REGION Network 2
   "TimeServerCom"(BatchEndTime := "OPC".CON_Material.NewBatchEndTime,
                   "Date" => "PrinterData".CON.PrinterBagData."Date",
                   "Time" => "PrinterData".CON.PrinterBagData."Time",
                   BatchStatus => "OPC".CON_Material.BatchStatus);
END_REGION

REGION Network 3
   IF NOT "PrinterData".CON.PrinterSelection THEN
       #Domino(RemoteAddress := "PrinterData".CON.PrinterBagData.RemoteAddress,   // "Domino_AX"
               ConnectionStatus := #ComandsSending_Domino.connected AND #BatchSending_Domino.connected,
               ID := 2,
               ConType := True,
               ArtFlag := #HandleComBag.ActualArtFlag,
               MDR_Flag := #HandleComBag.ActualMDR_Flag,
               BatchStatus := "OPC".CON_Material.BatchStatus,
               BatchNumber := "OPC".CON_Material.ActualBatchNumber,
               ArtBaseNumber := "OPC".CON_Material.ActualArtBaseNumber,
               MarketRegCode := "OPC".CON_Material.ActualMarketRegCode,
               ExtDate := "OPC".CON_Material.ActualBBD,
               "Date" := "PrinterData".CON.PrinterBagData."Date",
               "Time" := "PrinterData".CON.PrinterBagData."Time",
               PlainDataChanged := #HandleComBag.NewDataPlain,
               DataReceived := #ComandsSending_Domino.dataReceived,
               DataReceivedBatch := #BatchSending_Domino.dataReceived,
               DataSent := #ComandsSending_Domino.sending,
               DataSentBatch := #BatchSending_Domino.sending,
               TimeSynchPeriod := "TimeSynchPeriod",
               AlarmCheckPeriod := "AlarmCheckPeriod",
               RDataBatch := "PrinterData".CON.PrinterBagData.RdataBatch,
               RData := "PrinterData".CON.PrinterBagData.RData,
               NMDR_LabelName := "PrinterData".CON.PrinterBagData.NonMDR_LabelName,
               LabelSelecting := "PrinterData".CON.PrinterBagData.Initialization,
               ErrorIP => "CON_ErrorIP",
               BatchOK => "PrinterData".CON.PrinterBagData.BatchOK,
               TimeOK => "PrinterData".CON.PrinterBagData.TimeOK);
   END_IF;
END_REGION

REGION Network 4
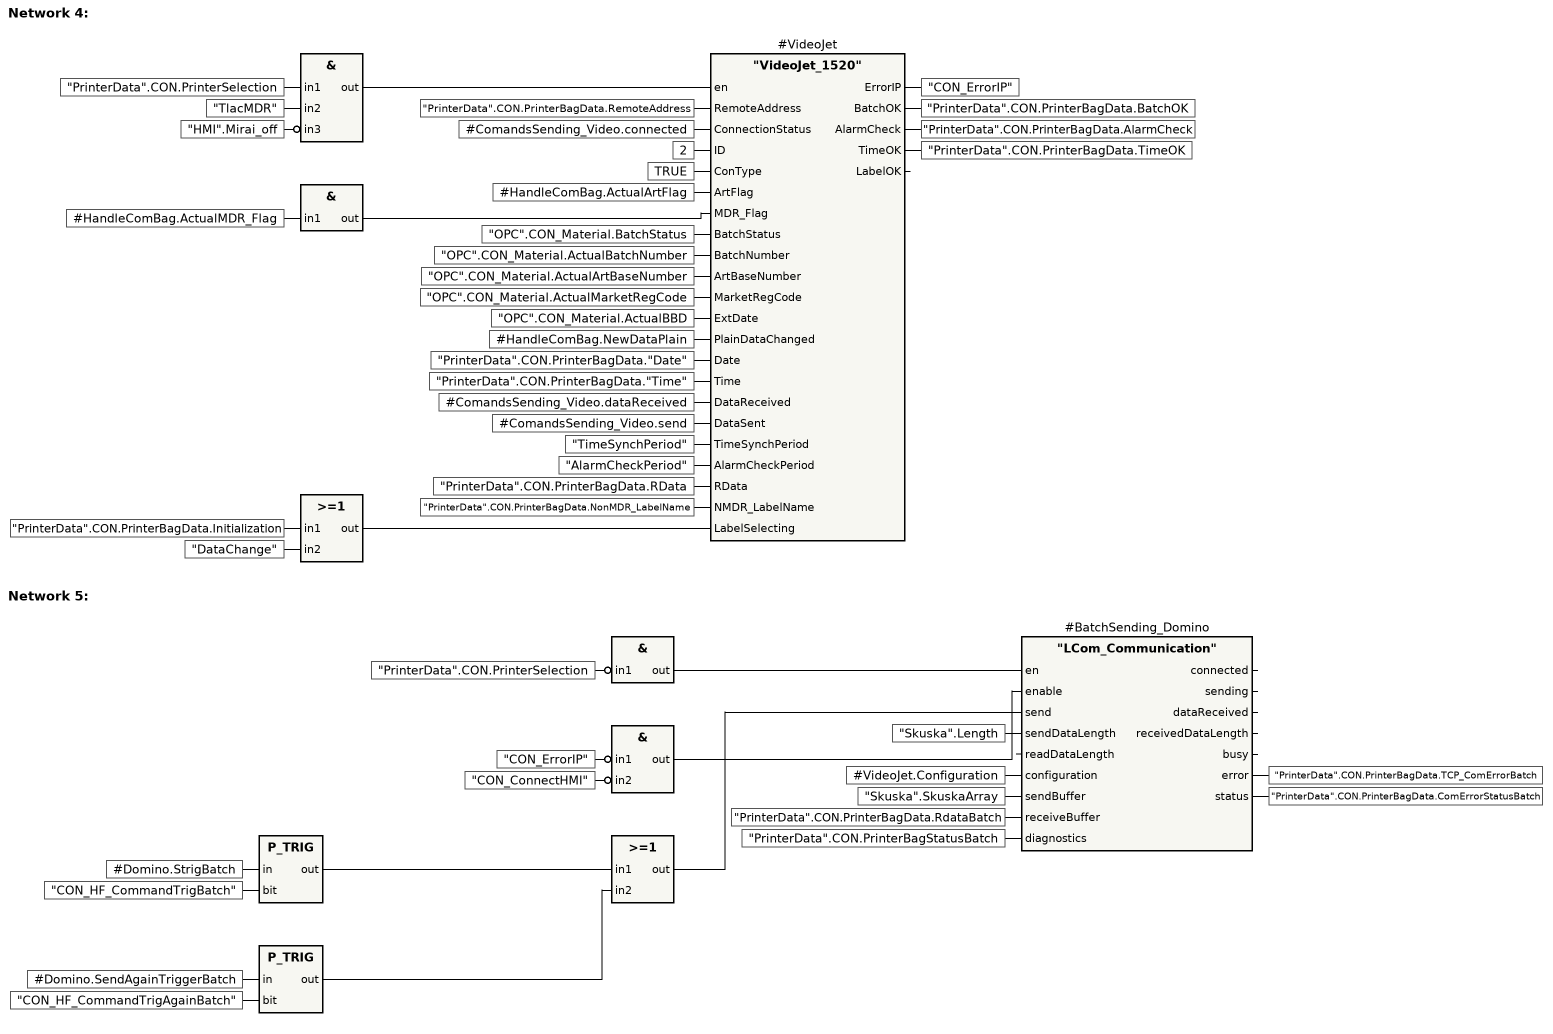
   IF "PrinterData".CON.PrinterSelection AND "TlacMDR" AND NOT "HMI".Mirai_off THEN
       #VideoJet(RemoteAddress := "PrinterData".CON.PrinterBagData.RemoteAddress,   // "VideoJet_1520"
                 ConnectionStatus := #ComandsSending_Video.connected,
                 ID := 2,
                 ConType := TRUE,
                 ArtFlag := #HandleComBag.ActualArtFlag,
                 MDR_Flag := #HandleComBag.ActualMDR_Flag,
                 BatchStatus := "OPC".CON_Material.BatchStatus,
                 BatchNumber := "OPC".CON_Material.ActualBatchNumber,
                 ArtBaseNumber := "OPC".CON_Material.ActualArtBaseNumber,
                 MarketRegCode := "OPC".CON_Material.ActualMarketRegCode,
                 ExtDate := "OPC".CON_Material.ActualBBD,
                 PlainDataChanged := #HandleComBag.NewDataPlain,
                 "Date" := "PrinterData".CON.PrinterBagData."Date",
                 "Time" := "PrinterData".CON.PrinterBagData."Time",
                 DataReceived := #ComandsSending_Video.dataReceived,
                 DataSent := #ComandsSending_Video.send,
                 TimeSynchPeriod := "TimeSynchPeriod",
                 AlarmCheckPeriod := "AlarmCheckPeriod",
                 RData := "PrinterData".CON.PrinterBagData.RData,
                 NMDR_LabelName := "PrinterData".CON.PrinterBagData.NonMDR_LabelName,
                 LabelSelecting := "PrinterData".CON.PrinterBagData.Initialization OR "DataChange",
                 ErrorIP => "CON_ErrorIP",
                 BatchOK => "PrinterData".CON.PrinterBagData.BatchOK,
                 AlarmCheck => "PrinterData".CON.PrinterBagData.AlarmCheck,
                 TimeOK => "PrinterData".CON.PrinterBagData.TimeOK);
   END_IF;
END_REGION

REGION Network 5
   #_w1 := #Domino.StrigBatch AND NOT "CON_HF_CommandTrigBatch";   // rising edge
   "CON_HF_CommandTrigBatch" := #Domino.StrigBatch;
   #_w2 := #Domino.SendAgainTriggerBatch AND NOT "CON_HF_CommandTrigAgainBatch";   // rising edge
   "CON_HF_CommandTrigAgainBatch" := #Domino.SendAgainTriggerBatch;
   IF NOT "PrinterData".CON.PrinterSelection THEN
       #BatchSending_Domino(enable := NOT "CON_ErrorIP" AND NOT "CON_ConnectHMI",   // "LCom_Communication"
                            send := #_w1 OR #_w2,
                            sendDataLength := "Skuska".Length,
                            configuration := #VideoJet.Configuration,
                            sendBuffer := "Skuska".SkuskaArray,
                            receiveBuffer := "PrinterData".CON.PrinterBagData.RdataBatch,
                            diagnostics := "PrinterData".CON.PrinterBagStatusBatch,
                            error => "PrinterData".CON.PrinterBagData.TCP_ComErrorBatch,
                            status => "PrinterData".CON.PrinterBagData.ComErrorStatusBatch);
   END_IF;
END_REGION

REGION Network 6
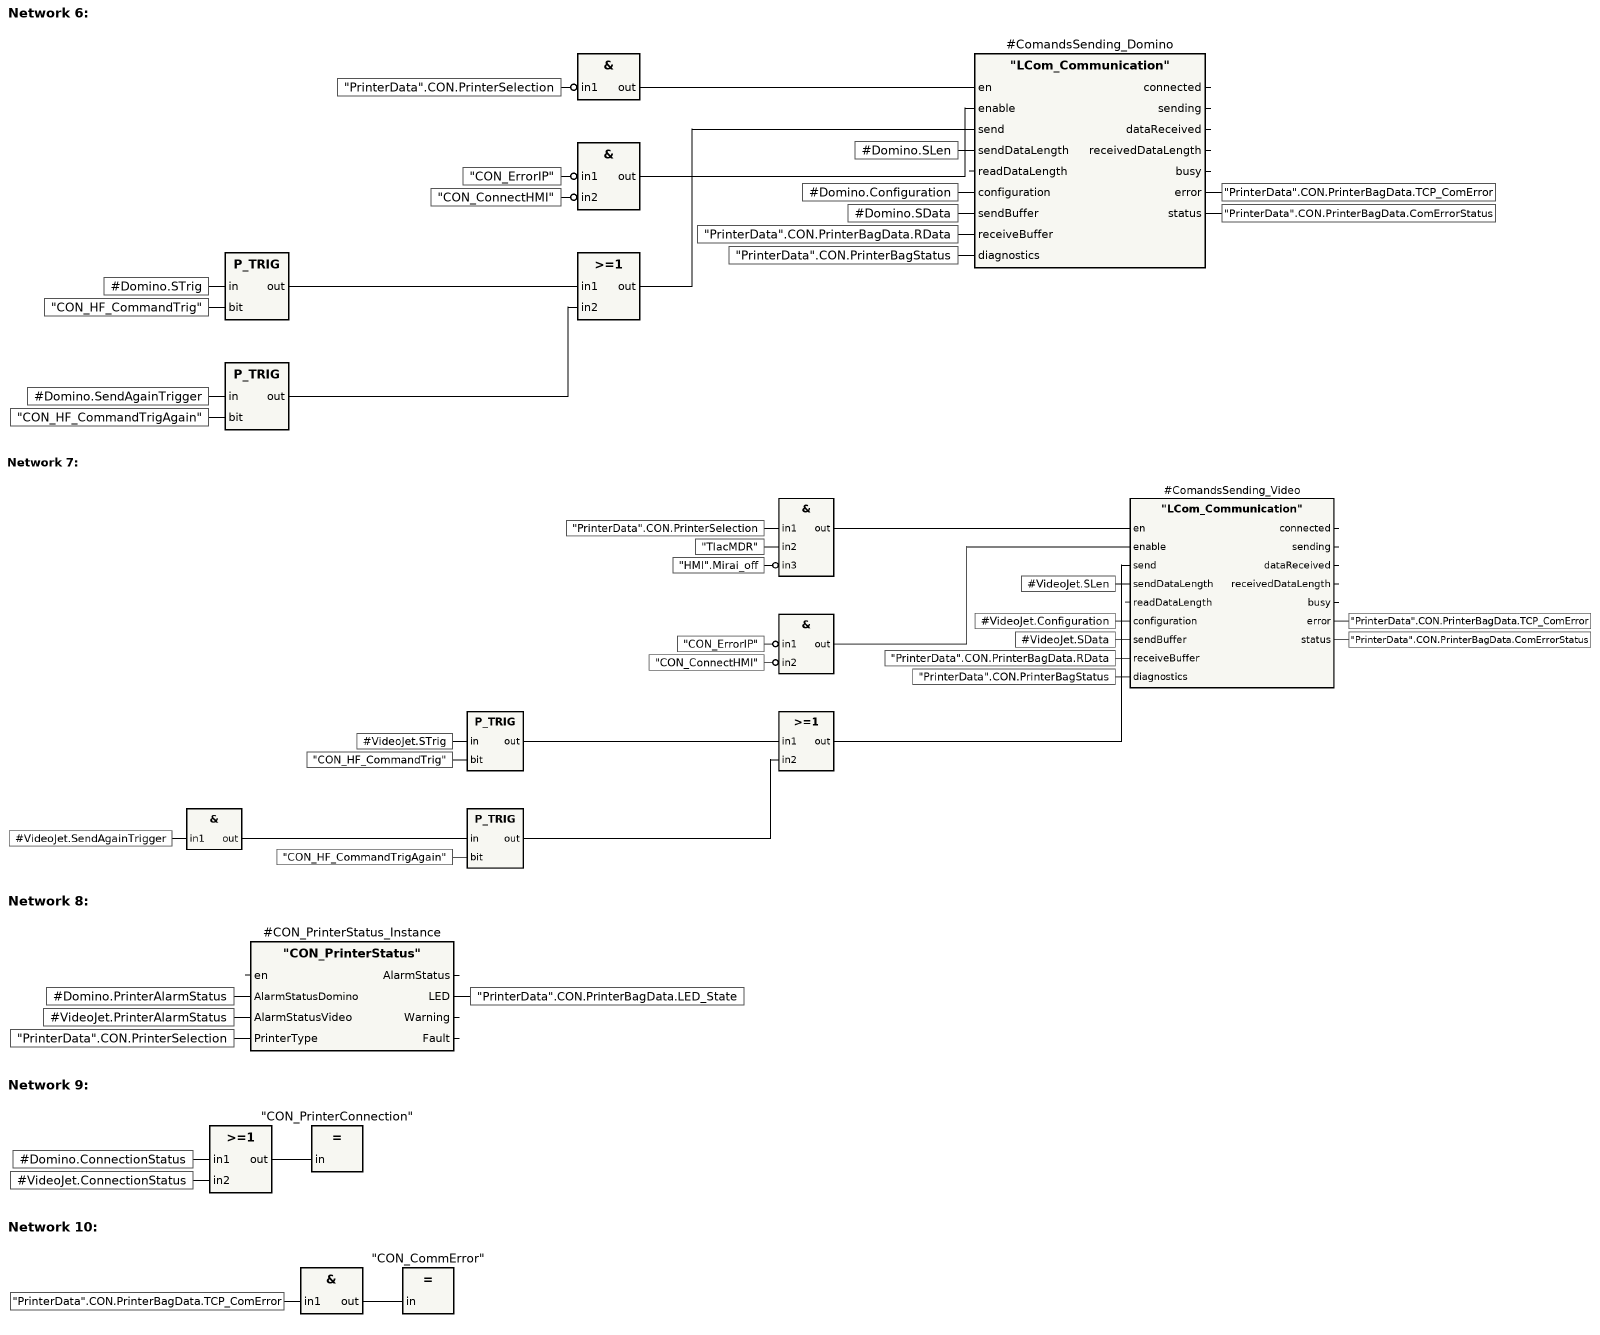
   #_w1 := #Domino.STrig AND NOT "CON_HF_CommandTrig";   // rising edge
   "CON_HF_CommandTrig" := #Domino.STrig;
   #_w2 := #Domino.SendAgainTrigger AND NOT "CON_HF_CommandTrigAgain";   // rising edge
   "CON_HF_CommandTrigAgain" := #Domino.SendAgainTrigger;
   IF NOT "PrinterData".CON.PrinterSelection THEN
       #ComandsSending_Domino(enable := NOT "CON_ErrorIP" AND NOT "CON_ConnectHMI",   // "LCom_Communication"
                              send := #_w1 OR #_w2,
                              sendDataLength := #Domino.SLen,
                              configuration := #Domino.Configuration,
                              sendBuffer := #Domino.SData,
                              receiveBuffer := "PrinterData".CON.PrinterBagData.RData,
                              diagnostics := "PrinterData".CON.PrinterBagStatus,
                              error => "PrinterData".CON.PrinterBagData.TCP_ComError,
                              status => "PrinterData".CON.PrinterBagData.ComErrorStatus);
   END_IF;
END_REGION

REGION Network 7
   #_w1 := #VideoJet.STrig AND NOT "CON_HF_CommandTrig";   // rising edge
   "CON_HF_CommandTrig" := #VideoJet.STrig;
   #_w2 := #VideoJet.SendAgainTrigger AND NOT "CON_HF_CommandTrigAgain";   // rising edge
   "CON_HF_CommandTrigAgain" := #VideoJet.SendAgainTrigger;
   IF "PrinterData".CON.PrinterSelection AND "TlacMDR" AND NOT "HMI".Mirai_off THEN
       #ComandsSending_Video(enable := NOT "CON_ErrorIP" AND NOT "CON_ConnectHMI",   // "LCom_Communication"
                             send := #_w1 OR #_w2,
                             sendDataLength := #VideoJet.SLen,
                             configuration := #VideoJet.Configuration,
                             sendBuffer := #VideoJet.SData,
                             receiveBuffer := "PrinterData".CON.PrinterBagData.RData,
                             diagnostics := "PrinterData".CON.PrinterBagStatus,
                             error => "PrinterData".CON.PrinterBagData.TCP_ComError,
                             status => "PrinterData".CON.PrinterBagData.ComErrorStatus);
   END_IF;
END_REGION

REGION Network 8
   #CON_PrinterStatus_Instance(AlarmStatusDomino := #Domino.PrinterAlarmStatus,   // "CON_PrinterStatus"
                           AlarmStatusVideo := #VideoJet.PrinterAlarmStatus,
                           PrinterType := "PrinterData".CON.PrinterSelection,
                           LED => "PrinterData".CON.PrinterBagData.LED_State);
END_REGION

REGION Network 9
   "CON_PrinterConnection" := #Domino.ConnectionStatus OR #VideoJet.ConnectionStatus;
END_REGION

REGION Network 10
   "CON_CommError" := "PrinterData".CON.PrinterBagData.TCP_ComError;
END_REGION
END_FUNCTION_BLOCK

FUNCTION_BLOCK "CON_PrinterStatus"   // FB14, FBD
{ S7_Optimized_Access := 'TRUE' }
VERSION : 0.1
   VAR_INPUT
      AlarmStatusDomino : Array[0..8] of Char;
      AlarmStatusVideo : Array[0..8] of Char;
      PrinterType : Bool;
   END_VAR
   VAR_OUTPUT
      AlarmStatus : String;
      LED : USInt;
      Warning : Bool;
      Fault : Bool;
   END_VAR
   VAR
      LEDStatus : String;
   END_VAR
BEGIN

REGION Network 1 (SCL)
   REGION led
       IF #PrinterType = FALSE THEN //Domino Printer
           Chars_TO_Strg(Chars := #AlarmStatusDomino,
                         pChars := 6,
                         Cnt := 2,
                         Strg => #LEDStatus);
           IF #LEDStatus = '00' OR #LEDStatus = '10' OR #LEDStatus = '01' THEN
               #LED := 3;
               #Warning := FALSE;
               #Fault := FALSE;
           ELSIF #LEDStatus = '02' OR #LEDStatus = '20' THEN
               #LED := 1;
               #Warning := TRUE;
               #Fault := FALSE;
           ELSIF #LEDStatus = '04' OR #LEDStatus = '40' THEN
               #LED := 2;
               #Warning := FALSE;
               #Fault := TRUE;
           ELSE
               #LED := 0;
               #Warning := FALSE;
               #Fault := FALSE;
           END_IF;
       ELSE //VideoJet Printer
           Chars_TO_Strg(Chars := #AlarmStatusVideo,
                         pChars := 7,
                         Cnt := 1,
                         Strg => #LEDStatus);
           IF #LEDStatus = '1' THEN
               #LED := 3;
               #Warning := FALSE;
               #Fault := FALSE;
           ELSIF #LEDStatus = '2' OR #LEDStatus = '3' THEN
               #LED := 1;
               #Warning := TRUE;
               #Fault := FALSE;
           ELSIF #LEDStatus = '4' THEN
               #LED := 2;
               #Warning := FALSE;
               #Fault := TRUE;
           ELSE
               #LED := 0;
               #Warning := FALSE;
               #Fault := FALSE;
           END_IF;
       END_IF;
   END_REGION
   REGION alarm
       //check the alarm
       IF #PrinterType = FALSE THEN //Domino Printer
           Chars_TO_Strg(Chars := #AlarmStatusDomino,
                         pChars := 3,
                         Cnt := 3,
                         Strg => #AlarmStatus);
           //IF Needed, create a conversion tabel to show the status of the printer       


       ELSE //VideoJet Printer
           Chars_TO_Strg(Chars := #AlarmStatusVideo,
                         pChars := 1,
                         Cnt := 6,
                         Strg => #AlarmStatus);
           //IF Needed, create a conversion tabel to show the status of the printer            


       END_IF;
   END_REGION
END_REGION
END_FUNCTION_BLOCK

FUNCTION_BLOCK "Reader_2D"   // FB15, LAD
{ S7_Optimized_Access := 'TRUE' }
VERSION : 0.1
   VAR_INPUT
      ExtTrigger : Bool;
      ResultAvailable : Bool;
      TriggerReady : Bool;
      TriggerAck : Bool;
      ResultID : Word;
      ResultCode : Word;
      ResultLength : Word;
      TriggerDelayTime : Time := T#10ms;
      SrcValue : ANY;
   END_VAR
   VAR_OUTPUT
      ID : UInt := 0;
      Flags : UInt := 0;
      Length : UInt := 0;
      TriggerEnable : Bool := false;
      TriggerReader : Bool := false;
      ResultsAck : Bool := false;
   END_VAR
   VAR_IN_OUT
      DstValue : ANY;
   END_VAR
   VAR
      T_DelayTrigger : TP_TIME;
      F_TRIG_Instance : F_TRIG;
      ResultPending : Bool;
      IntTrigger : Bool;
      HF_TriggerReader : Bool;
      HF_ResultsAck : Bool;
      IEC_Timer_0_Instance : TON_TIME;
      T_NoReadOutput : Bool;
   END_VAR
   VAR_TEMP
      BLKMOVRES : Int;
      Done : Bool;
   END_VAR
BEGIN

REGION Network 1 (SCL)
   REGION Triggering the camera 
       //Enable triggering via network 
       #TriggerEnable := TRUE;
       // intialize the triggering for determined delay time. 
     #T_DelayTrigger(IN:=#ExtTrigger,
                     PT:=#TriggerDelayTime);

    #F_TRIG_Instance(CLK:=#T_DelayTrigger.Q,
                     Q=>#IntTrigger);
    //if the conditions are met trigger the camera (If camera ready and trigger not already issued, issue trigger signal.)
    IF #TriggerReady = TRUE AND #ResultPending = FALSE AND #IntTrigger = TRUE AND #TriggerAck = FALSE AND #HF_TriggerReader = FALSE THEN
        #HF_TriggerReader := TRUE;
        #ResultPending := TRUE;
    END_IF;

    //Special CASE: IF results were already waiting before we issued a trigger, process those results instead OF issuing a new read sequence.
    IF #ResultAvailable = TRUE AND #ResultPending = FALSE THEN
        #ResultPending := TRUE;
    END_IF;
   END_REGION
   REGION Copy the data
       // Copy the data
       IF #ResultAvailable = TRUE AND #HF_ResultsAck = FALSE THEN
           #ID := #ResultID;
           #Flags := #ResultCode;
           #Length := #ResultLength;
           #BLKMOVRES := BLKMOV(SRCBLK := #SrcValue, DSTBLK => #DstValue);
           // act that the plc receive a results
           #HF_ResultsAck := TRUE;
       END_IF;
    //Reset trigger signal as soon as it is acknowledged
       IF #TriggerAck = TRUE AND #HF_ResultsAck = TRUE THEN
           #HF_TriggerReader := FALSE;
       END_IF;
    (*  Reset results acknowledge signal as soon as it is recognized BY the reader.
       This is the end OF the read sequence. Reset the "results pending" flag, set the
       output TO signal the operation is complete.
       Note, the reader signals "results acknowledge" BY setting "results available"
   TO zero.
       *)
       IF #HF_ResultsAck = TRUE AND #ResultAvailable = FALSE THEN
           #ResultPending := FALSE;
           #HF_ResultsAck := FALSE;
           #Done := True;
       END_IF;
     //  IF no read occurs within 90 seconds, cancel the read
     #IEC_Timer_0_Instance(IN:=#ResultPending,
                           PT:=T#90S,
                           Q=>#T_NoReadOutput);

     IF #T_NoReadOutput = TRUE THEN
         #HF_TriggerReader := FALSE;
         #HF_ResultsAck := FALSE;
         #ResultPending := FALSE;
         #Done := TRUE;
     END_IF;
     //assign the auxilary tags to the right ones
     #TriggerReader := #HF_TriggerReader;
     #ResultsAck:= #HF_ResultsAck;
   END_REGION
END_REGION
END_FUNCTION_BLOCK

FUNCTION_BLOCK "PlainHandle"   // FB16, LAD
{ S7_Optimized_Access := 'TRUE' }
VERSION : 0.1
   VAR_INPUT
      ResetFaults : Bool;
      NewBagDmcCode : String;
      NewBoxDmcCode : String;
      NewArticleNum : String;
      NewTotalInBag : String;
      NewTotalInBox : String;
      NewProductWeight : String;
      NewLineNumber : String;
      NewOrderNum : String;
   END_VAR
   VAR_OUTPUT
      LightAlarm : Bool;
      ActBagDmcCode : UDInt;
      ActBoxDmcCode : UDInt;
      ActArticleNum : String[12];
      ActTotalInBag : String[7];
      ActTotalInBox : String[7];
      ActProductWeight : String[10];
      ActLineNumber : String[5];
      ActOrderNum : String[12];
   END_VAR
   VAR_IN_OUT
      CommError : Bool;
      NoChange : Bool;
      NoData : Bool;
      DataChange : Bool;
   END_VAR
   VAR
      Aux1 : Bool;
      Aux0 : Bool;
      edge : Bool;
      CompareResult : Struct
         ResultBag : Bool;
         ResultBox : Bool;
         ResultArticleNUm : Bool;
         ResultTotalBag : Bool;
         ResultTotalBox : Bool;
         ResultWeight : Bool;
         ResultLineNumber : Bool;
         ResultOrderNum : Bool;
         PlainChange : Bool;
      END_STRUCT;
      OldCode : Struct
         DataDevice : String;
         BagDmcCode : String;
         BoxDmcCode : String;
         ArticleNum : String;
         TotalInBag : String;
         TotalInBox : String;
         ProductWeight : String;
         LineNumber : String;
         OrderNum : String;
      END_STRUCT;
      ActCode : Struct
         DataDevice : String;
         BagDmcCode : String;
         BoxDmcCode : String;
         ArticleNum : String;
         TotalInBag : String;
         TotalInBox : String;
         ProductWeight : String;
         LineNumber : String;
         OrderNum : String;
      END_STRUCT;
      CString : String := '                                                                               ';
      HeartBitNoPressent : Bool;
      PlainNoData : Bool;
      LiveBitTime : TON_TIME;
   END_VAR
   VAR_TEMP
      tmpI : Int;
   END_VAR
   VAR_TEMP   // added for the SCL form of the ladder/FBD networks
      _w1 : Bool;
   END_VAR
BEGIN

REGION Network 1
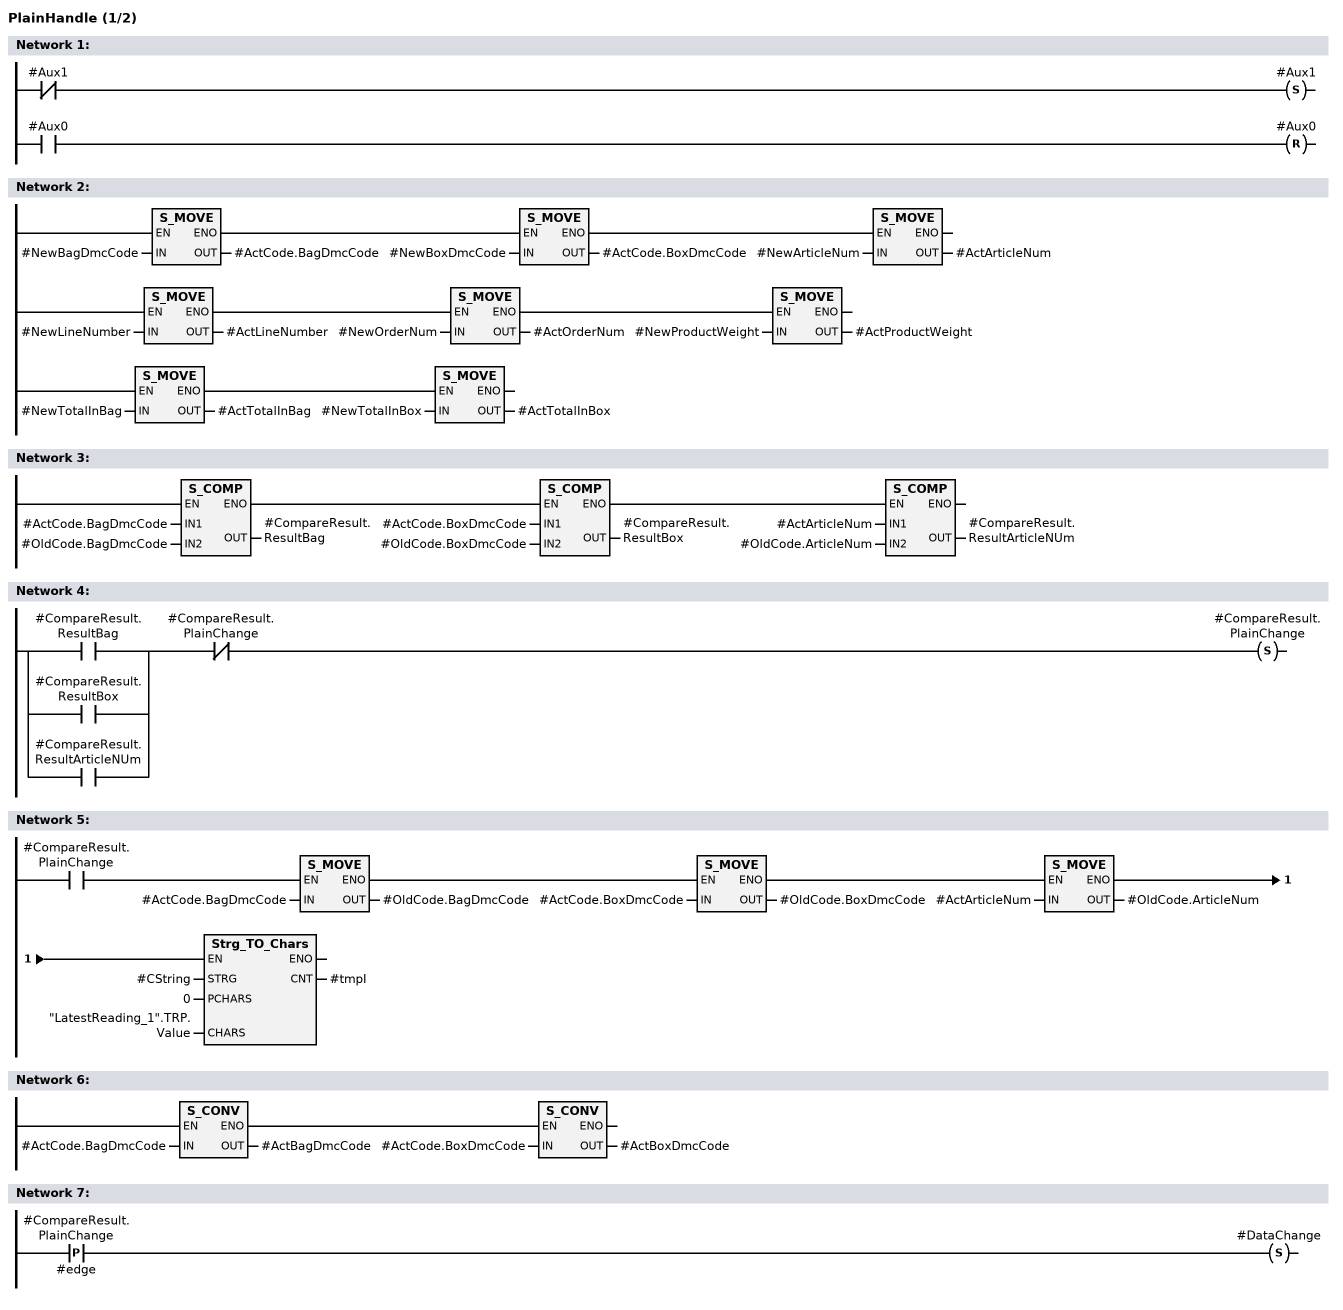
   RUNG wire#powerrail
      I_Contact( #Aux1 )
      S_Coil( #Aux1 )
   END_RUNG
   RUNG wire#powerrail
      Contact( #Aux0 )
      R_Coil( #Aux0 )
   END_RUNG
   // the same network as SCL:
   IF NOT #Aux1 THEN #Aux1 := TRUE; END_IF;
   IF #Aux0 THEN #Aux0 := FALSE; END_IF;
END_REGION

REGION Network 2
   RUNG wire#powerrail
      S_Move(in := #NewBagDmcCode, out => #ActCode.BagDmcCode)
      S_Move(in := #NewBoxDmcCode, out => #ActCode.BoxDmcCode)
      S_Move(in := #NewArticleNum, out => #ActArticleNum)
   END_RUNG
   RUNG wire#powerrail
      S_Move(in := #NewLineNumber, out => #ActLineNumber)
      S_Move(in := #NewOrderNum, out => #ActOrderNum)
      S_Move(in := #NewProductWeight, out => #ActProductWeight)
   END_RUNG
   RUNG wire#powerrail
      S_Move(in := #NewTotalInBag, out => #ActTotalInBag)
      S_Move(in := #NewTotalInBox, out => #ActTotalInBox)
   END_RUNG
   // the same network as SCL:
   #ActCode.BagDmcCode := #NewBagDmcCode;
   #ActCode.BoxDmcCode := #NewBoxDmcCode;
   #ActArticleNum := #NewArticleNum;
   #ActLineNumber := #NewLineNumber;
   #ActOrderNum := #NewOrderNum;
   #ActProductWeight := #NewProductWeight;
   #ActTotalInBag := #NewTotalInBag;
   #ActTotalInBox := #NewTotalInBox;
END_REGION

REGION Network 3
   // ENO of a box is taken as its EN; it also drops when the box reports an error
   S_COMP(IN1 := #ActCode.BagDmcCode, IN2 := #OldCode.BagDmcCode, OUT => #CompareResult.ResultBag);
   S_COMP(IN1 := #ActCode.BoxDmcCode, IN2 := #OldCode.BoxDmcCode, OUT => #CompareResult.ResultBox);
   S_COMP(IN1 := #ActArticleNum, IN2 := #OldCode.ArticleNum, OUT => #CompareResult.ResultArticleNUm);
END_REGION

REGION Network 4
   RUNG wire#powerrail
      Contact( #CompareResult.ResultBag )
      wire#w1
      I_Contact( #CompareResult.PlainChange )
      S_Coil( #CompareResult.PlainChange )
   END_RUNG
   RUNG wire#powerrail
      Contact( #CompareResult.ResultBox )
   END_RUNG wire#w1
   RUNG wire#powerrail
      Contact( #CompareResult.ResultArticleNUm )
   END_RUNG wire#w1
   // the same network as SCL:
   IF (#CompareResult.ResultBag OR #CompareResult.ResultBox OR #CompareResult.ResultArticleNUm) AND NOT #CompareResult.PlainChange THEN
       #CompareResult.PlainChange := TRUE;
   END_IF;
END_REGION

REGION Network 5
   // no SCL statement known for Strg_TO_Chars: written as a call
   IF #CompareResult.PlainChange THEN
       #OldCode.BagDmcCode := #ActCode.BagDmcCode;
       #OldCode.BoxDmcCode := #ActCode.BoxDmcCode;
       #OldCode.ArticleNum := #ActArticleNum;
       Strg_TO_Chars(Strg := #CString, pChars := 0, Chars := "LatestReading_1".TRP.Value, Cnt => #tmpI);
   END_IF;
END_REGION

REGION Network 6
   #ActBagDmcCode := S_CONV(IN := #ActCode.BagDmcCode);
   #ActBoxDmcCode := S_CONV(IN := #ActCode.BoxDmcCode);
END_REGION

REGION Network 7
   RUNG wire#powerrail
      P_Contact(operand := #CompareResult.PlainChange, bit := #edge)
      S_Coil( #DataChange )
   END_RUNG
   // the same network as SCL:
   #_w1 := #CompareResult.PlainChange AND NOT #edge;   // rising edge of #CompareResult.PlainChange
   #edge := #CompareResult.PlainChange;
   IF #_w1 THEN #DataChange := TRUE; END_IF;
END_REGION

REGION Network 8
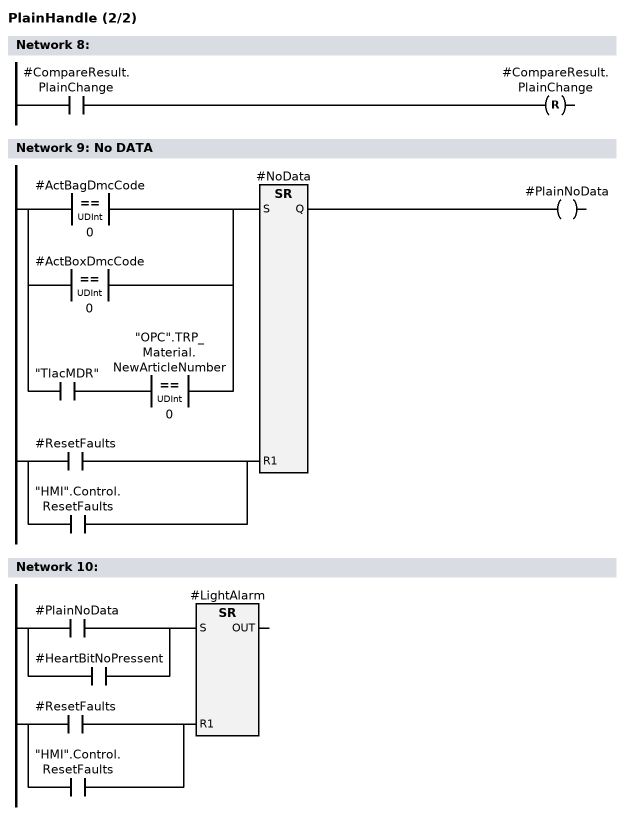
   RUNG wire#powerrail
      Contact( #CompareResult.PlainChange )
      R_Coil( #CompareResult.PlainChange )
   END_RUNG
   // the same network as SCL:
   IF #CompareResult.PlainChange THEN #CompareResult.PlainChange := FALSE; END_IF;
END_REGION

REGION Network 9: No DATA
   RUNG wire#powerrail
      { S7_Templates := "SrcType := UDInt" } EQ_Contact(in1 := #ActBagDmcCode, in2 := 0)
      wire#w1
      S_SR(operand := #NoData, r1 := wire#w2)
      Coil( #PlainNoData )
   END_RUNG
   RUNG wire#powerrail
      { S7_Templates := "SrcType := UDInt" } EQ_Contact(in1 := #ActBoxDmcCode, in2 := 0)
   END_RUNG wire#w1
   RUNG wire#powerrail
      Contact( "TlacMDR" )
      { S7_Templates := "SrcType := UDInt" } EQ_Contact(in1 := "OPC".TRP_Material.NewArticleNumber, in2 := 0)
   END_RUNG wire#w1
   RUNG wire#powerrail
      Contact( #ResetFaults )
   END_RUNG wire#w2
   RUNG wire#powerrail
      Contact( "HMI".Control.ResetFaults )
   END_RUNG wire#w2
   // the same network as SCL:
   IF (#ActBagDmcCode = 0) OR (#ActBoxDmcCode = 0) OR ("TlacMDR" AND ("OPC".TRP_Material.NewArticleNumber = 0)) THEN
       #NoData := TRUE;   // SR flip-flop
   END_IF;
   IF #ResetFaults OR "HMI".Control.ResetFaults THEN #NoData := FALSE; END_IF;
   #PlainNoData := #NoData;
END_REGION

REGION Network 10
   RUNG wire#powerrail
      Contact( #PlainNoData )
      wire#w1
      S_SR(operand := #LightAlarm, r1 := wire#w2)
   END_RUNG
   RUNG wire#powerrail
      Contact( #HeartBitNoPressent )
   END_RUNG wire#w1
   RUNG wire#powerrail
      Contact( #ResetFaults )
   END_RUNG wire#w2
   RUNG wire#powerrail
      Contact( "HMI".Control.ResetFaults )
   END_RUNG wire#w2
   // the same network as SCL:
   IF #PlainNoData OR #HeartBitNoPressent THEN
       #LightAlarm := TRUE;   // SR flip-flop
   END_IF;
   IF #ResetFaults OR "HMI".Control.ResetFaults THEN #LightAlarm := FALSE; END_IF;
END_REGION
END_FUNCTION_BLOCK

FUNCTION_BLOCK "TRP_PrinterStatus"   // FB17, FBD
{ S7_Optimized_Access := 'TRUE' }
VERSION : 0.1
   VAR_INPUT
      PrinterStatus : Array[0..31] of Bool;
      PrinterConnection : Bool;
   END_VAR
   VAR_OUTPUT
      TRP_ErrorsW1 : Word;
      TRP_ErrorsW2 : Word;
      LED : USInt;
   END_VAR
   VAR
      AlarmDataW1 : Word;
      AlamsBits1 AT AlarmDataW1 : Array[0..15] of Bool;
      AlarmDataW2 : Word;
      AlarmBits2 AT AlarmDataW2 : Array[0..15] of Bool;
   END_VAR
   VAR_TEMP
      i : Int;
   END_VAR
BEGIN

REGION Network 1 (SCL)
   REGION alarm
     //will be complete 
       FOR #i:=0 TO 15 DO
           #AlamsBits1[#i] := #PrinterStatus[#i];
       END_FOR;
       FOR #i:=16 TO 31 DO
           #AlarmBits2[#i-16] := #PrinterStatus[#i];
       END_FOR;
       #TRP_ErrorsW1 := #AlarmDataW1;
       #TRP_ErrorsW2 := #AlarmDataW2;
   END_REGION
   REGION led
       // Led of the printer. 
       IF #AlarmDataW1 = 0 AND #AlarmDataW2 = 0 AND #PrinterConnection = 1 THEN
           #LED := 0; //ready to print
       ELSE
           #LED := 2; //fault or warning
       END_IF;
   END_REGION
END_REGION
END_FUNCTION_BLOCK

FUNCTION_BLOCK "ReaderVerification"   // FB18, FBD
{ S7_Optimized_Access := 'TRUE' }
VERSION : 0.1
   VAR_INPUT
      Decoded : Array[0..79] of Char;
      BatchNumber : String;
      GTIN_Number : String;
      ArtNumber : String;
      MachineID : String;
      "Date" : String;
      ExtDate : String;
      ReaderRead : Bool;
      ReaderNoRead : Bool;
      ExtTrigger : Bool;
      ResetFaults : Bool;
      ResetCounters : Bool;
   END_VAR
   VAR_OUTPUT
      MisMatchFault : Bool;
      NoReadFault : Bool;
      TriggerFault : Bool;
   END_VAR
   VAR_IN_OUT
      NumGross : UDInt;
      NumRead : UDInt;
      NumNoRead : UDInt;
      NumMatch : UDInt;
      NumMisMatch : UDInt;
   END_VAR
   VAR
      ReadTimer : TP_TIME;
      NoReadTimer : TP_TIME;
      DecodedBatch : String;
      DecodedGTIN : String;
      DecodedArticle : String;
      DecodedTime : String;
      DecodedMachine : String;
      DecodedCounter : String;
      DecodedDate : String;
      DecodedExt : String;
   END_VAR
   VAR RETAIN
      MatchC : CTU_INT;
      Match : Bool;
   END_VAR
   VAR
      MisMatch : Bool;
      ValidDataF : F_TRIG;
   END_VAR
   VAR RETAIN
      NoReadCounter : CTU_INT;
      TriggerCounterNoRead : CTU_INT;
   END_VAR
   VAR
      WatchDog : TON_TIME;
      ExtTriggerR : R_TRIG;
      ReaderReadR : R_TRIG;
      ReaderNoReadR : R_TRIG;
   END_VAR
   VAR RETAIN
      TriggerCounterMischMatch : CTU_INT;
   END_VAR
   VAR_TEMP
      ResetDummy : Bool;
      WatchDogActive : Bool;
      NoReadActive : Bool;
   END_VAR
   VAR CONSTANT
      TimeRead : Time := T#60ms;
      TimeNoRead : Time := T#500ms;
      TimeTrigger : Time := T#1M;
      GTIN_P : USInt := 2;
      BatchP : USInt := 18;
      ArticleP : USInt := 31;
      TimeP : USInt := 44;
      MachineP : USInt := 50;
      CounterP : USInt := 53;
      DateP : USInt := 61;
      ExtP : USInt := 69;
      TriggersMaxNoRead : USInt := 100;
      NoReadLimit : USInt := 3;
   END_VAR
BEGIN

REGION Network 1 (SCL)
   REGION Decoded data
       // process the decod data
       Chars_TO_Strg(Chars := #Decoded,
                     pChars := #GTIN_P,
                     Cnt := 14,
                     Strg => #DecodedGTIN);
       Chars_TO_Strg(Chars:=#Decoded,
                     pChars:=#BatchP,
                     Cnt:=10,
                     Strg=>#DecodedBatch);
       Chars_TO_Strg(Chars:=#Decoded,
                     pChars:=#ArticleP,
                     Cnt:=10,
                     Strg=>#DecodedArticle);
      Chars_TO_Strg(Chars:=#Decoded,
                    pChars:=#TimeP,
                    Cnt:=6,
                    Strg=>#DecodedTime);
       Chars_TO_Strg(Chars:=#Decoded,
                     pChars:=#MachineP,
                     Cnt:=3,
                     Strg=>#DecodedMachine);
     Chars_TO_Strg(Chars:=#Decoded,
                   pChars:=#CounterP,
                   Cnt:=5,
                   Strg=>#DecodedCounter);
     Chars_TO_Strg(Chars := #Decoded,
                   pChars := #DateP,
                   Cnt := 6,
                   Strg => #DecodedDate);
     Chars_TO_Strg(Chars := #Decoded,
                   pChars := #ExtP,
                   Cnt := 6,
                   Strg => #DecodedExt
     );
     IF #DecodedExt = 'XXXXXX' OR #DecodedExt = '      ' THEN
         #DecodedExt := '';
     END_IF;
   END_REGION
   REGION CameraOutput
       //Make sure to activate outputs in the reader 
       #ReadTimer(IN := #ReaderRead,
                  PT := #TimeRead);
       #NoReadTimer(IN := #ReaderNoRead,
                    PT := #TimeNoRead);
       #ValidDataF(CLK := #ReadTimer.Q); //wait for data to be ready

       IF #ValidDataF.Q = TRUE THEN // reader has a good read and the data is valid for processitng
           IF #DecodedGTIN = #GTIN_Number AND #DecodedBatch = #BatchNumber AND #DecodedArticle = #ArtNumber  AND #DecodedExt = #ExtDate THEN
               #Match := TRUE;
               #MisMatch := FALSE;
           ELSE
               IF #DecodedGTIN <> 'XXXXXXXXXXXXXX' THEN
                   #Match := FALSE;
                   #MisMatch := TRUE;
               END_IF;
           END_IF;
       ELSE
           #Match := FALSE;
           #MisMatch := FALSE;
       END_IF;
   END_REGION
   REGION Fault
       //MisMatch Fault
       #TriggerCounterMischMatch( CU := #MisMatch,
                                 R := #ResetFaults OR #Match,
                                 PV := #NoReadLimit,
                                  Q => #MisMatchFault);

       //count 100 product (3 no read per 100)
       #TriggerCounterNoRead(CU := #ExtTrigger,
                             R := #ResetDummy,
                             PV := #TriggersMaxNoRead);
       IF #TriggerCounterNoRead.CV >= #TriggersMaxNoRead THEN
           #ResetDummy := TRUE;
       ELSE
           #ResetDummy := FALSE;
       END_IF;
       //NoRead Fault
       #NoReadCounter(CU := #ReaderNoRead OR (#ReaderRead AND #DecodedGTIN = 'XXXXXXXXXXXXXX'),
                      R := #ResetFaults OR #TriggerCounterNoRead.QU,
                      PV := #NoReadLimit,
                      Q => #NoReadActive);
       IF #NoReadActive = TRUE AND #ResetFaults = FALSE THEN
           #NoReadFault := TRUE;
       END_IF;
       #WatchDog(IN := #ExtTrigger,
                 PT := #TimeTrigger,
                 Q => #WatchDogActive);
       IF #WatchDogActive = TRUE AND #ResetFaults = FALSE THEN
           #TriggerFault := TRUE;
       END_IF;
       //Reset the Faults
       IF #ResetFaults = TRUE THEN
           #NoReadFault := FALSE;
           #MisMatchFault := FALSE;
           #TriggerFault := FALSE;
       END_IF;
   END_REGION

   REGION Count
   //detect positive edge on input
   #ExtTriggerR(CLK:=#ExtTrigger);
   #ReaderReadR(CLK:=#ReaderRead);
   #ReaderNoReadR(CLK := #ReaderNoRead OR (#ValidDataF.Q = TRUE AND #ReaderRead AND #DecodedGTIN = 'XXXXXXXXXXXXXX'));
       IF #ExtTriggerR.Q = TRUE THEN
           "Counter_32Bit_1"(Varia := 1,
                           CountedValue := #NumGross);
       END_IF;
       IF #ReaderReadR.Q = TRUE THEN
           "Counter_32Bit_1"(Varia := 1,
                           CountedValue := #NumRead);
       END_IF;
       IF #ReaderNoReadR.Q = TRUE THEN
           "Counter_32Bit_1"(Varia := 1,
                           CountedValue := #NumNoRead);
       END_IF;
       IF #ValidDataF.Q = TRUE AND #Match = TRUE THEN
           "Counter_32Bit_1"(Varia := 1,
                           CountedValue := #NumMatch);
       END_IF;
       IF #ValidDataF.Q = TRUE AND #MisMatch = TRUE THEN
           "Counter_32Bit_1"(Varia := 1,
                           CountedValue := #NumMisMatch);
       END_IF;
       IF #ResetCounters = TRUE THEN
           #NumGross := 0;
           #NumNoRead := 0;
           #NumRead := 0;
           #NumMatch := 0;
           #NumMisMatch := 0;
           #TriggerCounterNoRead.CV := 0;
       END_IF;
   END_REGION
END_REGION
END_FUNCTION_BLOCK

FUNCTION_BLOCK "HandleCom"   // FB20, FBD
{ S7_Optimized_Access := 'TRUE' }
VERSION : 0.1
   VAR_INPUT
      NewMaterialNumber : UDInt;
   END_VAR
   VAR_OUTPUT
      ArticleChange : Bool;
   END_VAR
   VAR_IN_OUT
      ActualMaterialNumber : UDInt;
   END_VAR
   VAR_TEMP
      i : Int;
   END_VAR
BEGIN

REGION Network 1
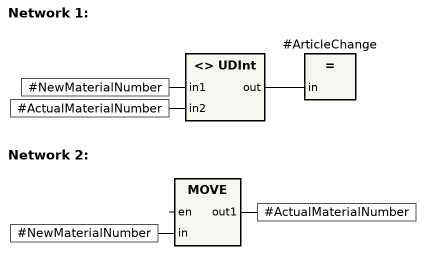
   #ArticleChange := #NewMaterialNumber <> #ActualMaterialNumber;
END_REGION

REGION Network 2
   #ActualMaterialNumber := #NewMaterialNumber;
END_REGION
END_FUNCTION_BLOCK

FUNCTION_BLOCK "TRP_PlainHandle"   // FB22, FBD
{ S7_Optimized_Access := 'TRUE' }
VERSION : 0.1
   VAR_INPUT
      NewGTIN_Num : String;
      NewBatchNum : String;
      NewArtNum : UDInt;
      NewMatchineID : String;
      NewBBD : String;
   END_VAR
   VAR_OUTPUT
      ActualGTIN_NumSTR : String;
      ActualBatchNumSTR : String;
      ActualArtNumSTR : String;
      ActualMachineID_STR : String;
      ActualBBD_STR : String;
   END_VAR
   VAR
      PlainDataChange : Bool;
      ExtDateChange : Bool;
      ActualGTIN_Num : String;
      ActualBatchNum : String;
      ActualArtNum : UDInt;
      ActualMachineID : String;
      ActualExtDate : String;
   END_VAR
   VAR_TEMP
      NewGTIN_Len : UInt;
      NewBatchLen : UInt;
      NewMachinID_Len : UInt;
      Correction : Array[0..13] of Char;
      CorrectionSTR : String;
      i : Int;
      Dummy1 : UInt;
      ArtSTR : String;
      NewArtSTR : String;
      ArtChar : Array[0..9] of Char;
      MachineIDChar : Array[0..4] of Char;
   END_VAR
   VAR CONSTANT
      GTIN_Size : UInt := 14;
      BatchSize : UInt := 10;
      ArtSize : UInt := 10;
      MachineID_Size : UInt := 3;
   END_VAR
BEGIN

REGION Network 1 (SCL)
   REGION batch changing
       // check for input data changing
       IF #NewGTIN_Num <> #ActualGTIN_Num OR #NewBatchNum <> #ActualBatchNum OR #NewArtNum <>#ActualArtNum OR #NewBBD <> #ActualExtDate OR #NewMatchineID <> #ActualMachineID THEN
           #PlainDataChange  := TRUE;
       ELSE
           #PlainDataChange := FALSE;
       END_IF;
       IF #NewBBD <> #ActualExtDate OR #NewArtNum <> #ActualArtNum THEN
           #ExtDateChange := TRUE;
       ELSE
           #ExtDateChange := FALSE;
       END_IF;
   END_REGION
   REGION assign new data 
       FOR #i := 0 TO 13 DO
           #Correction[#i] := '0';
       END_FOR;
       // save a copy of variables coming from plain to check the changes
       #ActualGTIN_Num := #NewGTIN_Num;
       #ActualBatchNum := #NewBatchNum;
       #ActualArtNum := #NewArtNum;
       #ActualMachineID := #NewMatchineID;
       #ActualExtDate := #NewBBD;
       //check the size of variables and prepare them for printing
       //Actual GTIN in 14
       #NewGTIN_Len := INT_TO_UINT(LEN(#NewGTIN_Num));
       IF #NewGTIN_Len < #GTIN_Size  THEN
          Chars_TO_Strg(Chars:=#Correction,
                        pChars:=0,
                        Cnt:=(#GTIN_Size -#NewGTIN_Len),
                        Strg=>#CorrectionSTR);
          #ActualGTIN_NumSTR:= CONCAT(IN1:=#CorrectionSTR, IN2:=#NewGTIN_Num);
      ELSE
          #ActualGTIN_NumSTR := #NewGTIN_Num;
      END_IF;
      //Actual Batch in 10 digits (3 factoryID+7 batch ID)
      #NewBatchLen := INT_TO_UINT(LEN(#NewBatchNum));
      IF #NewBatchLen < #BatchSize THEN
          Chars_TO_Strg(Chars := #Correction,
                        pChars := 0,
                        Cnt := (#BatchSize - #NewBatchLen),
                        Strg => #CorrectionSTR);
          #ActualBatchNumSTR := CONCAT(IN1 := #CorrectionSTR, IN2 := #NewBatchNum);
      ELSE
          #ActualBatchNumSTR := #NewBatchNum;
      END_IF;
      //Actual Article number in 10 
      VAL_STRG(IN:=#NewArtNum,
               SIZE:=UINT_TO_USINT(#ArtSize),
               PREC:=0,
               FORMAT:=0,
               P:=1,
               OUT=>#ArtSTR);
   Strg_TO_Chars(Strg:=#ArtSTR,
                 pChars:=0,
                 Cnt=>#Dummy1,
                 Chars:=#ArtChar);
   FOR #i := 0 TO UINT_TO_INT(#ArtSize-1) DO
       IF #ArtChar[#i] = ' ' THEN
           #ArtChar[#i] := '0';
       END_IF;
   END_FOR;
   Chars_TO_Strg(Chars:=#ArtChar,
                 pChars:=0,
                 Cnt:=#ArtSize,
                 Strg=>#NewArtSTR);
   #ActualArtNumSTR := #NewArtSTR;
     //take the 3 digits out of 5 for the machine ID 
   #NewMachinID_Len := INT_TO_UINT(LEN(#NewMatchineID));
   IF #NewMachinID_Len > #MachineID_Size THEN
       Strg_TO_Chars(Strg := #NewMatchineID,
                     pChars := 0,
                     Cnt => #Dummy1,
                     Chars := #MachineIDChar);
       Chars_TO_Strg(Chars := #MachineIDChar,
                     pChars := 2,
                     Cnt := #MachineID_Size,
                     Strg => #ActualMachineID_STR);
   ELSIF #NewMachinID_Len <#MachineID_Size THEN
       #ActualMachineID_STR := '000';
   ELSE
       #ActualMachineID_STR := #NewMatchineID;
   END_IF;
   //Actual Expiration date in 6
   #ActualBBD_STR := #NewBBD;
   END_REGION
END_REGION
END_FUNCTION_BLOCK

